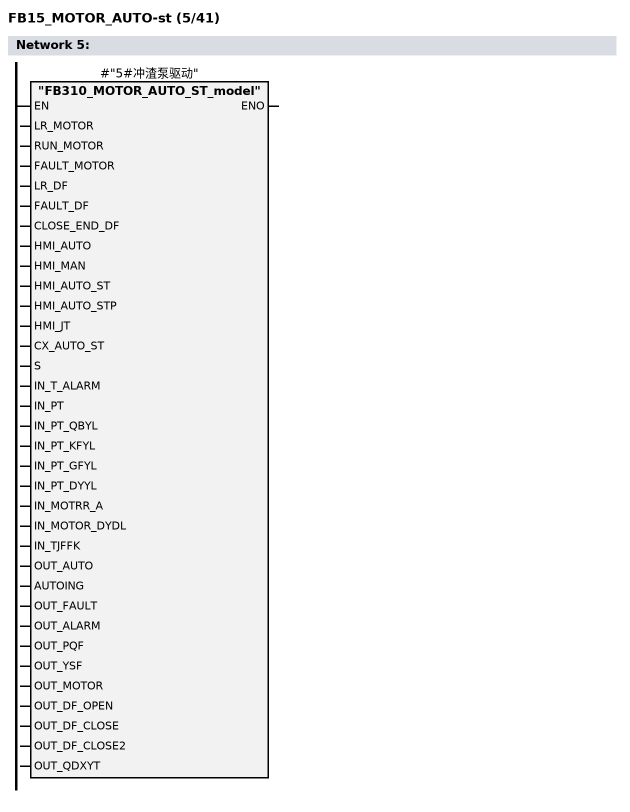
   RUNG wire#powerrail
      #"5#冲渣泵驱动"(LR_MOTOR :=, RUN_MOTOR :=, FAULT_MOTOR :=, LR_DF :=, FAULT_DF :=, CLOSE_END_DF :=, HMI_AUTO :=, HMI_MAN :=, HMI_AUTO_ST :=, HMI_AUTO_STP :=, HMI_JT :=, CX_AUTO_ST :=, S :=, IN_T_ALARM :=, IN_PT :=, IN_PT_QBYL :=, IN_PT_KFYL :=, IN_PT_GFYL :=, IN_PT_DYYL :=, IN_MOTRR_A :=, IN_MOTOR_DYDL :=, IN_TJFFK :=, OUT_AUTO :=, AUTOING :=, OUT_FAULT :=, OUT_ALARM :=, OUT_PQF :=, OUT_YSF :=, OUT_MOTOR :=, OUT_DF_OPEN :=, OUT_DF_CLOSE :=, OUT_DF_CLOSE2 :=, OUT_QDXYT :=)
   END_RUNG
   // the same network as SCL:
   #"5#冲渣泵驱动"();   // "FB310_MOTOR_AUTO_ST_model"
END_REGION

REGION Network 6
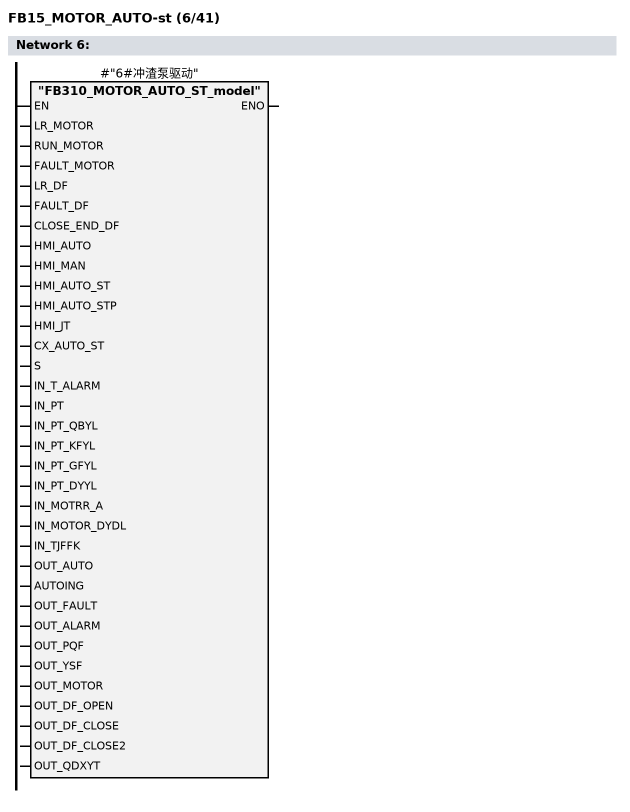
   RUNG wire#powerrail
      #"6#冲渣泵驱动"(LR_MOTOR :=, RUN_MOTOR :=, FAULT_MOTOR :=, LR_DF :=, FAULT_DF :=, CLOSE_END_DF :=, HMI_AUTO :=, HMI_MAN :=, HMI_AUTO_ST :=, HMI_AUTO_STP :=, HMI_JT :=, CX_AUTO_ST :=, S :=, IN_T_ALARM :=, IN_PT :=, IN_PT_QBYL :=, IN_PT_KFYL :=, IN_PT_GFYL :=, IN_PT_DYYL :=, IN_MOTRR_A :=, IN_MOTOR_DYDL :=, IN_TJFFK :=, OUT_AUTO :=, AUTOING :=, OUT_FAULT :=, OUT_ALARM :=, OUT_PQF :=, OUT_YSF :=, OUT_MOTOR :=, OUT_DF_OPEN :=, OUT_DF_CLOSE :=, OUT_DF_CLOSE2 :=, OUT_QDXYT :=)
   END_RUNG
   // the same network as SCL:
   #"6#冲渣泵驱动"();   // "FB310_MOTOR_AUTO_ST_model"
END_REGION

REGION Network 7
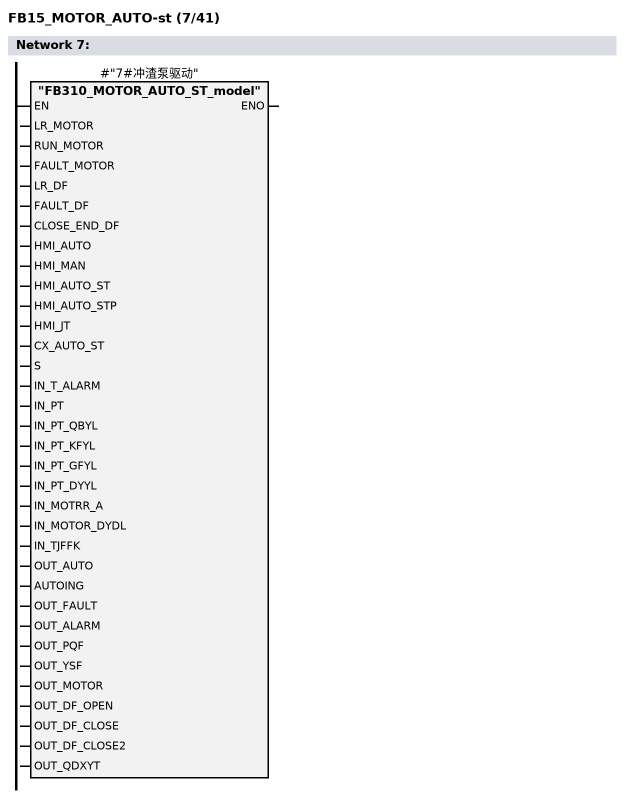
   RUNG wire#powerrail
      #"7#冲渣泵驱动"(LR_MOTOR :=, RUN_MOTOR :=, FAULT_MOTOR :=, LR_DF :=, FAULT_DF :=, CLOSE_END_DF :=, HMI_AUTO :=, HMI_MAN :=, HMI_AUTO_ST :=, HMI_AUTO_STP :=, HMI_JT :=, CX_AUTO_ST :=, S :=, IN_T_ALARM :=, IN_PT :=, IN_PT_QBYL :=, IN_PT_KFYL :=, IN_PT_GFYL :=, IN_PT_DYYL :=, IN_MOTRR_A :=, IN_MOTOR_DYDL :=, IN_TJFFK :=, OUT_AUTO :=, AUTOING :=, OUT_FAULT :=, OUT_ALARM :=, OUT_PQF :=, OUT_YSF :=, OUT_MOTOR :=, OUT_DF_OPEN :=, OUT_DF_CLOSE :=, OUT_DF_CLOSE2 :=, OUT_QDXYT :=)
   END_RUNG
   // the same network as SCL:
   #"7#冲渣泵驱动"();   // "FB310_MOTOR_AUTO_ST_model"
END_REGION

REGION Network 8
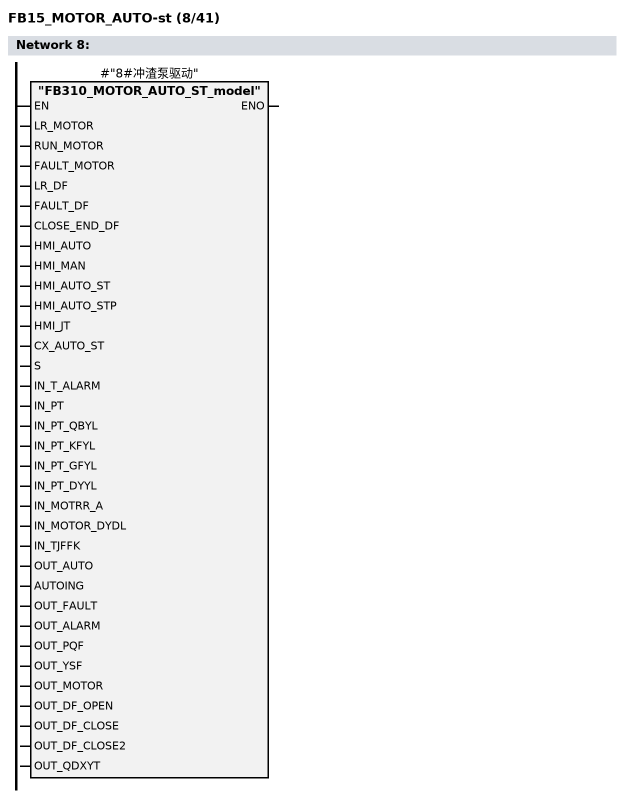
   RUNG wire#powerrail
      #"8#冲渣泵驱动"(LR_MOTOR :=, RUN_MOTOR :=, FAULT_MOTOR :=, LR_DF :=, FAULT_DF :=, CLOSE_END_DF :=, HMI_AUTO :=, HMI_MAN :=, HMI_AUTO_ST :=, HMI_AUTO_STP :=, HMI_JT :=, CX_AUTO_ST :=, S :=, IN_T_ALARM :=, IN_PT :=, IN_PT_QBYL :=, IN_PT_KFYL :=, IN_PT_GFYL :=, IN_PT_DYYL :=, IN_MOTRR_A :=, IN_MOTOR_DYDL :=, IN_TJFFK :=, OUT_AUTO :=, AUTOING :=, OUT_FAULT :=, OUT_ALARM :=, OUT_PQF :=, OUT_YSF :=, OUT_MOTOR :=, OUT_DF_OPEN :=, OUT_DF_CLOSE :=, OUT_DF_CLOSE2 :=, OUT_QDXYT :=)
   END_RUNG
   // the same network as SCL:
   #"8#冲渣泵驱动"();   // "FB310_MOTOR_AUTO_ST_model"
END_REGION

REGION Network 9
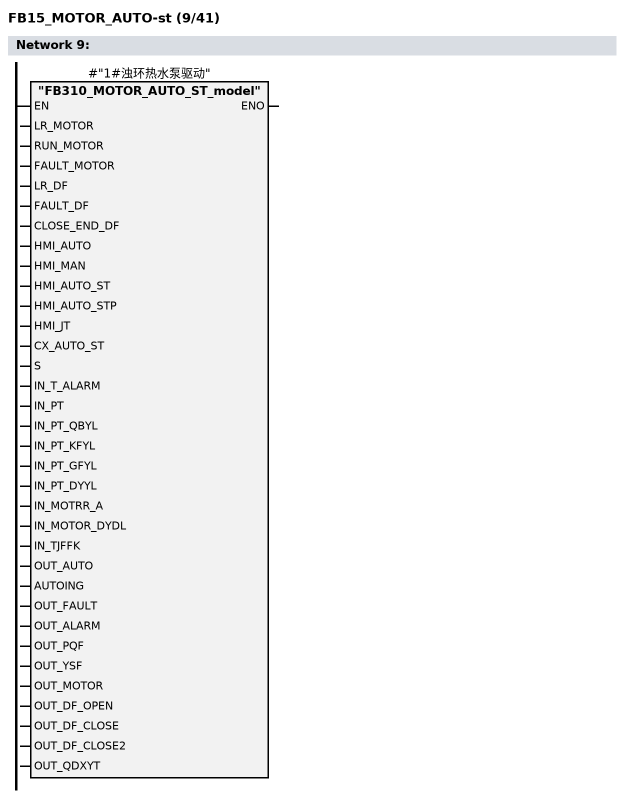
   RUNG wire#powerrail
      #"1#浊环热水泵驱动"(LR_MOTOR :=, RUN_MOTOR :=, FAULT_MOTOR :=, LR_DF :=, FAULT_DF :=, CLOSE_END_DF :=, HMI_AUTO :=, HMI_MAN :=, HMI_AUTO_ST :=, HMI_AUTO_STP :=, HMI_JT :=, CX_AUTO_ST :=, S :=, IN_T_ALARM :=, IN_PT :=, IN_PT_QBYL :=, IN_PT_KFYL :=, IN_PT_GFYL :=, IN_PT_DYYL :=, IN_MOTRR_A :=, IN_MOTOR_DYDL :=, IN_TJFFK :=, OUT_AUTO :=, AUTOING :=, OUT_FAULT :=, OUT_ALARM :=, OUT_PQF :=, OUT_YSF :=, OUT_MOTOR :=, OUT_DF_OPEN :=, OUT_DF_CLOSE :=, OUT_DF_CLOSE2 :=, OUT_QDXYT :=)
   END_RUNG
   // the same network as SCL:
   #"1#浊环热水泵驱动"();   // "FB310_MOTOR_AUTO_ST_model"
END_REGION

REGION Network 10
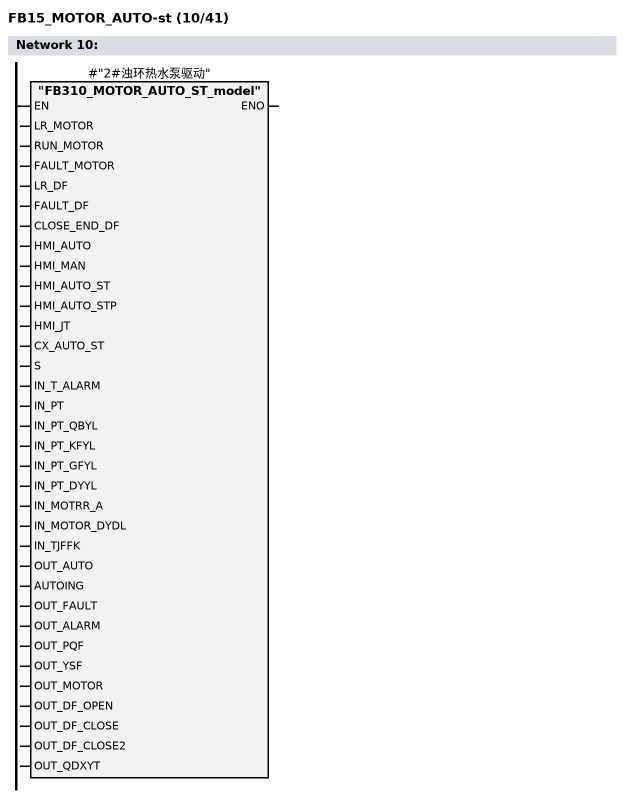
   RUNG wire#powerrail
      #"2#浊环热水泵驱动"(LR_MOTOR :=, RUN_MOTOR :=, FAULT_MOTOR :=, LR_DF :=, FAULT_DF :=, CLOSE_END_DF :=, HMI_AUTO :=, HMI_MAN :=, HMI_AUTO_ST :=, HMI_AUTO_STP :=, HMI_JT :=, CX_AUTO_ST :=, S :=, IN_T_ALARM :=, IN_PT :=, IN_PT_QBYL :=, IN_PT_KFYL :=, IN_PT_GFYL :=, IN_PT_DYYL :=, IN_MOTRR_A :=, IN_MOTOR_DYDL :=, IN_TJFFK :=, OUT_AUTO :=, AUTOING :=, OUT_FAULT :=, OUT_ALARM :=, OUT_PQF :=, OUT_YSF :=, OUT_MOTOR :=, OUT_DF_OPEN :=, OUT_DF_CLOSE :=, OUT_DF_CLOSE2 :=, OUT_QDXYT :=)
   END_RUNG
   // the same network as SCL:
   #"2#浊环热水泵驱动"();   // "FB310_MOTOR_AUTO_ST_model"
END_REGION

REGION Network 11
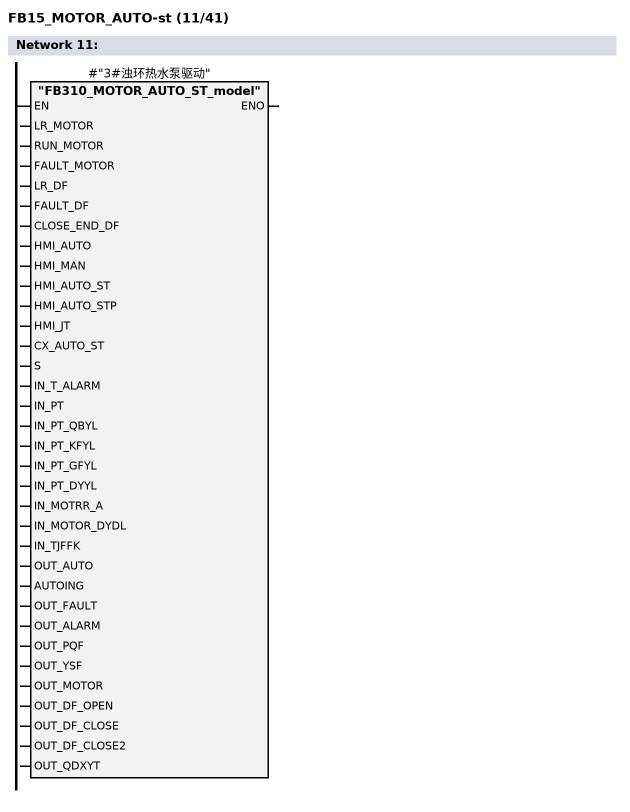
   RUNG wire#powerrail
      #"3#浊环热水泵驱动"(LR_MOTOR :=, RUN_MOTOR :=, FAULT_MOTOR :=, LR_DF :=, FAULT_DF :=, CLOSE_END_DF :=, HMI_AUTO :=, HMI_MAN :=, HMI_AUTO_ST :=, HMI_AUTO_STP :=, HMI_JT :=, CX_AUTO_ST :=, S :=, IN_T_ALARM :=, IN_PT :=, IN_PT_QBYL :=, IN_PT_KFYL :=, IN_PT_GFYL :=, IN_PT_DYYL :=, IN_MOTRR_A :=, IN_MOTOR_DYDL :=, IN_TJFFK :=, OUT_AUTO :=, AUTOING :=, OUT_FAULT :=, OUT_ALARM :=, OUT_PQF :=, OUT_YSF :=, OUT_MOTOR :=, OUT_DF_OPEN :=, OUT_DF_CLOSE :=, OUT_DF_CLOSE2 :=, OUT_QDXYT :=)
   END_RUNG
   // the same network as SCL:
   #"3#浊环热水泵驱动"();   // "FB310_MOTOR_AUTO_ST_model"
END_REGION

REGION Network 12
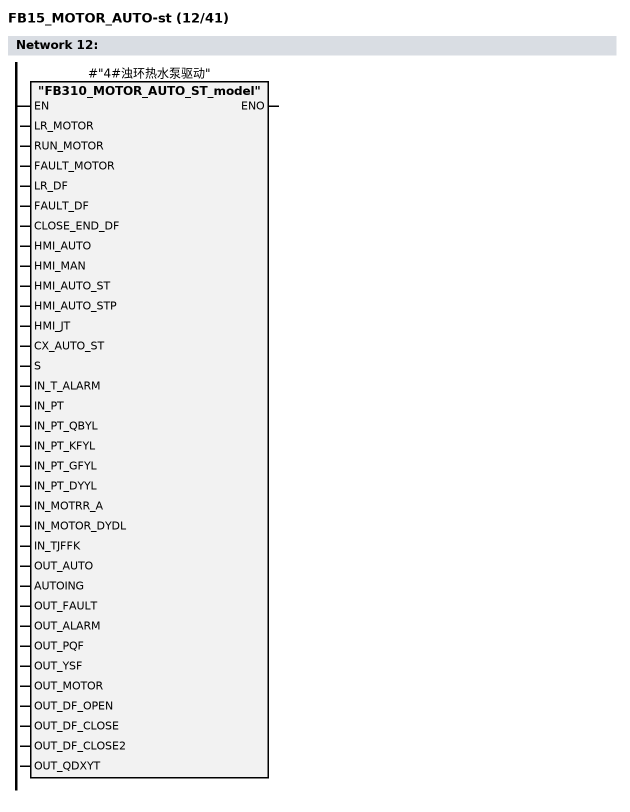
   RUNG wire#powerrail
      #"4#浊环热水泵驱动"(LR_MOTOR :=, RUN_MOTOR :=, FAULT_MOTOR :=, LR_DF :=, FAULT_DF :=, CLOSE_END_DF :=, HMI_AUTO :=, HMI_MAN :=, HMI_AUTO_ST :=, HMI_AUTO_STP :=, HMI_JT :=, CX_AUTO_ST :=, S :=, IN_T_ALARM :=, IN_PT :=, IN_PT_QBYL :=, IN_PT_KFYL :=, IN_PT_GFYL :=, IN_PT_DYYL :=, IN_MOTRR_A :=, IN_MOTOR_DYDL :=, IN_TJFFK :=, OUT_AUTO :=, AUTOING :=, OUT_FAULT :=, OUT_ALARM :=, OUT_PQF :=, OUT_YSF :=, OUT_MOTOR :=, OUT_DF_OPEN :=, OUT_DF_CLOSE :=, OUT_DF_CLOSE2 :=, OUT_QDXYT :=)
   END_RUNG
   // the same network as SCL:
   #"4#浊环热水泵驱动"();   // "FB310_MOTOR_AUTO_ST_model"
END_REGION

REGION Network 13
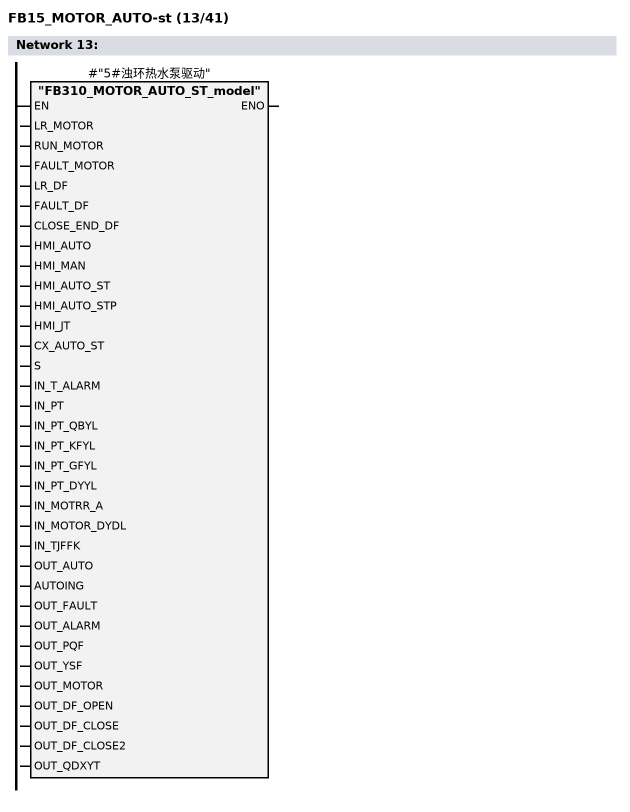
   RUNG wire#powerrail
      #"5#浊环热水泵驱动"(LR_MOTOR :=, RUN_MOTOR :=, FAULT_MOTOR :=, LR_DF :=, FAULT_DF :=, CLOSE_END_DF :=, HMI_AUTO :=, HMI_MAN :=, HMI_AUTO_ST :=, HMI_AUTO_STP :=, HMI_JT :=, CX_AUTO_ST :=, S :=, IN_T_ALARM :=, IN_PT :=, IN_PT_QBYL :=, IN_PT_KFYL :=, IN_PT_GFYL :=, IN_PT_DYYL :=, IN_MOTRR_A :=, IN_MOTOR_DYDL :=, IN_TJFFK :=, OUT_AUTO :=, AUTOING :=, OUT_FAULT :=, OUT_ALARM :=, OUT_PQF :=, OUT_YSF :=, OUT_MOTOR :=, OUT_DF_OPEN :=, OUT_DF_CLOSE :=, OUT_DF_CLOSE2 :=, OUT_QDXYT :=)
   END_RUNG
   // the same network as SCL:
   #"5#浊环热水泵驱动"();   // "FB310_MOTOR_AUTO_ST_model"
END_REGION

REGION Network 14
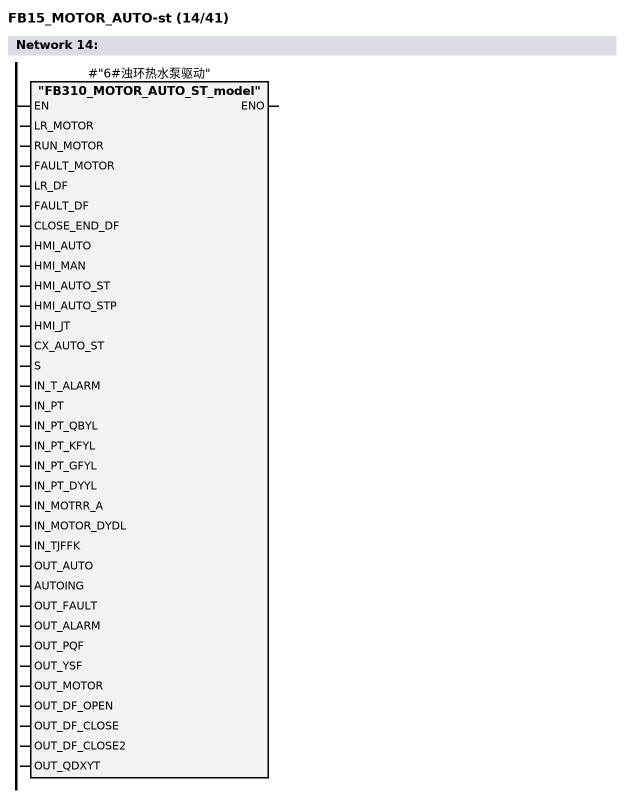
   RUNG wire#powerrail
      #"6#浊环热水泵驱动"(LR_MOTOR :=, RUN_MOTOR :=, FAULT_MOTOR :=, LR_DF :=, FAULT_DF :=, CLOSE_END_DF :=, HMI_AUTO :=, HMI_MAN :=, HMI_AUTO_ST :=, HMI_AUTO_STP :=, HMI_JT :=, CX_AUTO_ST :=, S :=, IN_T_ALARM :=, IN_PT :=, IN_PT_QBYL :=, IN_PT_KFYL :=, IN_PT_GFYL :=, IN_PT_DYYL :=, IN_MOTRR_A :=, IN_MOTOR_DYDL :=, IN_TJFFK :=, OUT_AUTO :=, AUTOING :=, OUT_FAULT :=, OUT_ALARM :=, OUT_PQF :=, OUT_YSF :=, OUT_MOTOR :=, OUT_DF_OPEN :=, OUT_DF_CLOSE :=, OUT_DF_CLOSE2 :=, OUT_QDXYT :=)
   END_RUNG
   // the same network as SCL:
   #"6#浊环热水泵驱动"();   // "FB310_MOTOR_AUTO_ST_model"
END_REGION

REGION Network 15
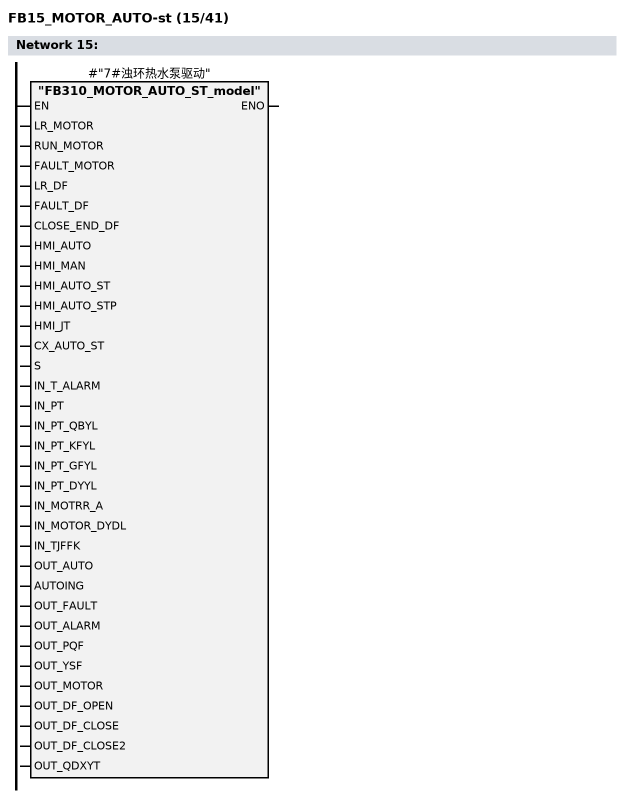
   RUNG wire#powerrail
      #"7#浊环热水泵驱动"(LR_MOTOR :=, RUN_MOTOR :=, FAULT_MOTOR :=, LR_DF :=, FAULT_DF :=, CLOSE_END_DF :=, HMI_AUTO :=, HMI_MAN :=, HMI_AUTO_ST :=, HMI_AUTO_STP :=, HMI_JT :=, CX_AUTO_ST :=, S :=, IN_T_ALARM :=, IN_PT :=, IN_PT_QBYL :=, IN_PT_KFYL :=, IN_PT_GFYL :=, IN_PT_DYYL :=, IN_MOTRR_A :=, IN_MOTOR_DYDL :=, IN_TJFFK :=, OUT_AUTO :=, AUTOING :=, OUT_FAULT :=, OUT_ALARM :=, OUT_PQF :=, OUT_YSF :=, OUT_MOTOR :=, OUT_DF_OPEN :=, OUT_DF_CLOSE :=, OUT_DF_CLOSE2 :=, OUT_QDXYT :=)
   END_RUNG
   // the same network as SCL:
   #"7#浊环热水泵驱动"();   // "FB310_MOTOR_AUTO_ST_model"
END_REGION

REGION Network 16
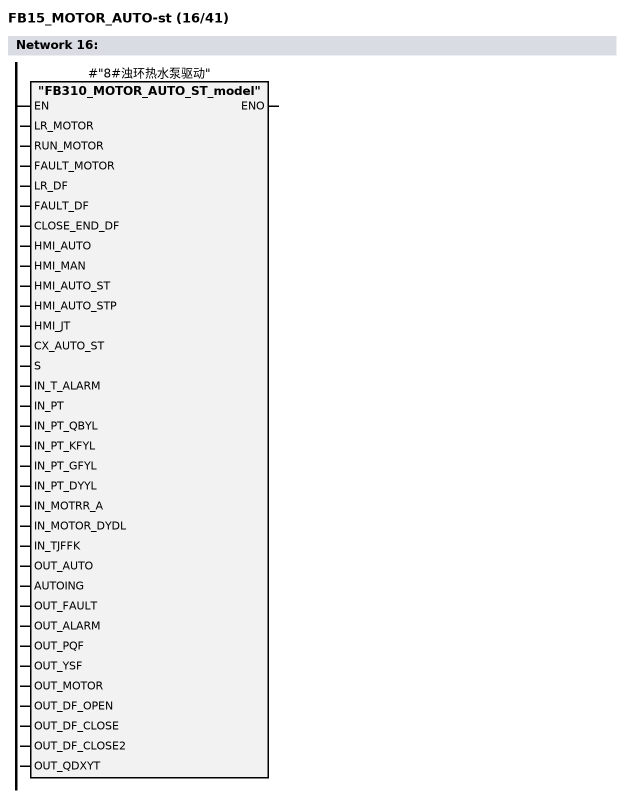
   RUNG wire#powerrail
      #"8#浊环热水泵驱动"(LR_MOTOR :=, RUN_MOTOR :=, FAULT_MOTOR :=, LR_DF :=, FAULT_DF :=, CLOSE_END_DF :=, HMI_AUTO :=, HMI_MAN :=, HMI_AUTO_ST :=, HMI_AUTO_STP :=, HMI_JT :=, CX_AUTO_ST :=, S :=, IN_T_ALARM :=, IN_PT :=, IN_PT_QBYL :=, IN_PT_KFYL :=, IN_PT_GFYL :=, IN_PT_DYYL :=, IN_MOTRR_A :=, IN_MOTOR_DYDL :=, IN_TJFFK :=, OUT_AUTO :=, AUTOING :=, OUT_FAULT :=, OUT_ALARM :=, OUT_PQF :=, OUT_YSF :=, OUT_MOTOR :=, OUT_DF_OPEN :=, OUT_DF_CLOSE :=, OUT_DF_CLOSE2 :=, OUT_QDXYT :=)
   END_RUNG
   // the same network as SCL:
   #"8#浊环热水泵驱动"();   // "FB310_MOTOR_AUTO_ST_model"
END_REGION

REGION Network 17
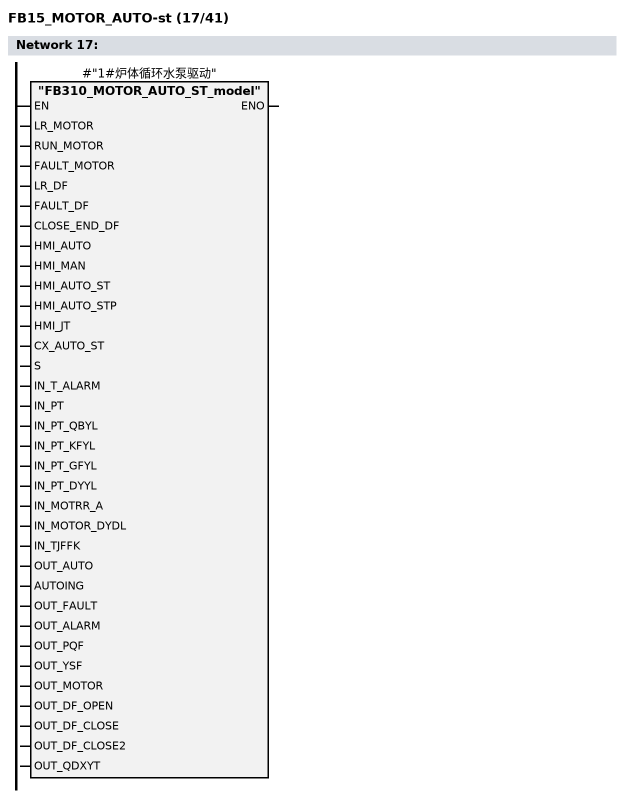
   RUNG wire#powerrail
      #"1#炉体循环水泵驱动"(LR_MOTOR :=, RUN_MOTOR :=, FAULT_MOTOR :=, LR_DF :=, FAULT_DF :=, CLOSE_END_DF :=, HMI_AUTO :=, HMI_MAN :=, HMI_AUTO_ST :=, HMI_AUTO_STP :=, HMI_JT :=, CX_AUTO_ST :=, S :=, IN_T_ALARM :=, IN_PT :=, IN_PT_QBYL :=, IN_PT_KFYL :=, IN_PT_GFYL :=, IN_PT_DYYL :=, IN_MOTRR_A :=, IN_MOTOR_DYDL :=, IN_TJFFK :=, OUT_AUTO :=, AUTOING :=, OUT_FAULT :=, OUT_ALARM :=, OUT_PQF :=, OUT_YSF :=, OUT_MOTOR :=, OUT_DF_OPEN :=, OUT_DF_CLOSE :=, OUT_DF_CLOSE2 :=, OUT_QDXYT :=)
   END_RUNG
   // the same network as SCL:
   #"1#炉体循环水泵驱动"();   // "FB310_MOTOR_AUTO_ST_model"
END_REGION

REGION Network 18
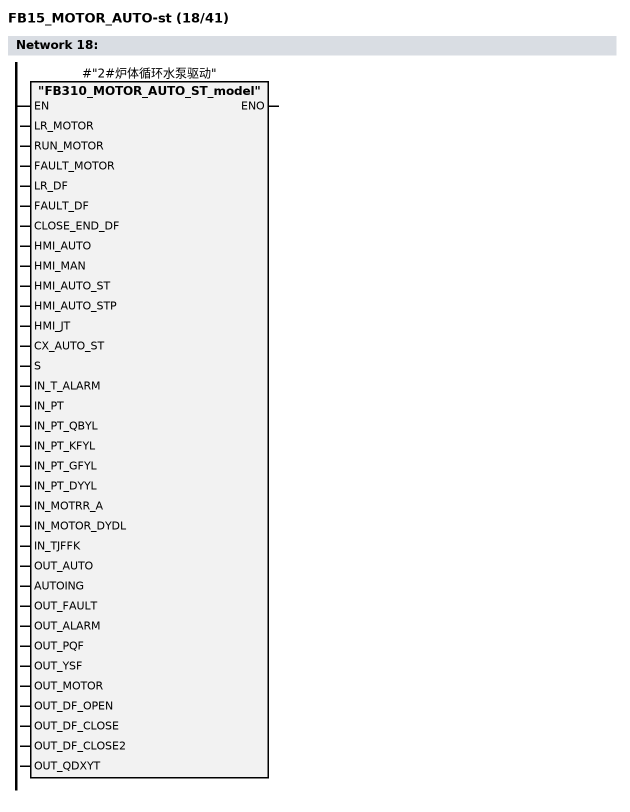
   RUNG wire#powerrail
      #"2#炉体循环水泵驱动"(LR_MOTOR :=, RUN_MOTOR :=, FAULT_MOTOR :=, LR_DF :=, FAULT_DF :=, CLOSE_END_DF :=, HMI_AUTO :=, HMI_MAN :=, HMI_AUTO_ST :=, HMI_AUTO_STP :=, HMI_JT :=, CX_AUTO_ST :=, S :=, IN_T_ALARM :=, IN_PT :=, IN_PT_QBYL :=, IN_PT_KFYL :=, IN_PT_GFYL :=, IN_PT_DYYL :=, IN_MOTRR_A :=, IN_MOTOR_DYDL :=, IN_TJFFK :=, OUT_AUTO :=, AUTOING :=, OUT_FAULT :=, OUT_ALARM :=, OUT_PQF :=, OUT_YSF :=, OUT_MOTOR :=, OUT_DF_OPEN :=, OUT_DF_CLOSE :=, OUT_DF_CLOSE2 :=, OUT_QDXYT :=)
   END_RUNG
   // the same network as SCL:
   #"2#炉体循环水泵驱动"();   // "FB310_MOTOR_AUTO_ST_model"
END_REGION

REGION Network 19
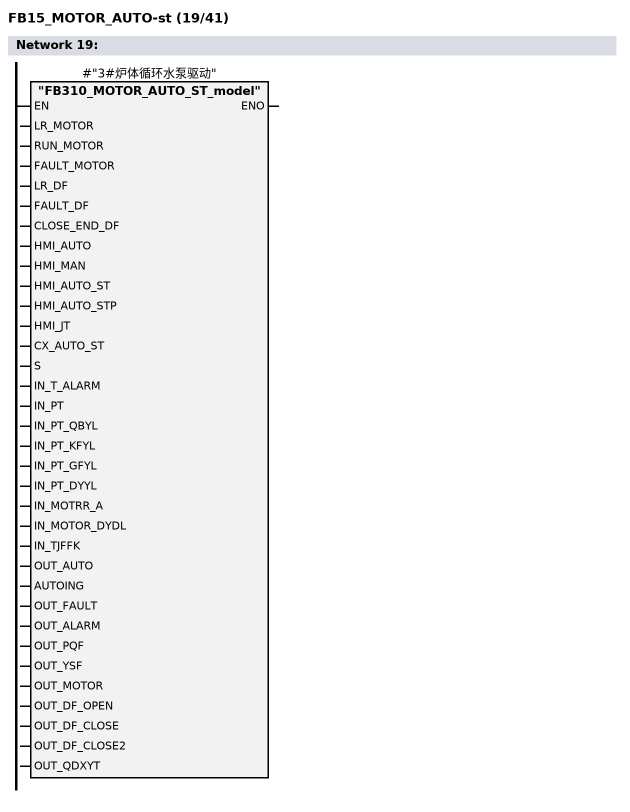
   RUNG wire#powerrail
      #"3#炉体循环水泵驱动"(LR_MOTOR :=, RUN_MOTOR :=, FAULT_MOTOR :=, LR_DF :=, FAULT_DF :=, CLOSE_END_DF :=, HMI_AUTO :=, HMI_MAN :=, HMI_AUTO_ST :=, HMI_AUTO_STP :=, HMI_JT :=, CX_AUTO_ST :=, S :=, IN_T_ALARM :=, IN_PT :=, IN_PT_QBYL :=, IN_PT_KFYL :=, IN_PT_GFYL :=, IN_PT_DYYL :=, IN_MOTRR_A :=, IN_MOTOR_DYDL :=, IN_TJFFK :=, OUT_AUTO :=, AUTOING :=, OUT_FAULT :=, OUT_ALARM :=, OUT_PQF :=, OUT_YSF :=, OUT_MOTOR :=, OUT_DF_OPEN :=, OUT_DF_CLOSE :=, OUT_DF_CLOSE2 :=, OUT_QDXYT :=)
   END_RUNG
   // the same network as SCL:
   #"3#炉体循环水泵驱动"();   // "FB310_MOTOR_AUTO_ST_model"
END_REGION

REGION Network 20
